           // Increment the actual configured devices, store the state and
           // HW_ID as an numerical value (UINT)
           #statActualConfiguredDevices := #statActualConfiguredDevices + 1;
         ELSE
           ;
         END_IF;

       ELSE
         ; // Device not configured
       END_IF;
     END_FOR;

     #ioSystemData.actualConfiguredDevices := #statActualConfiguredDevices;

     // Mark parameter "Next Device" of the last device in the list
     // --> "Next Device" = negative --> Last device in the list
     #ioSystemData.devices[#statLastDevice].nextDevice := #LAST_DEVICE;

   END_IF; // New IO System detected at input

   #ioSystemData.error := FALSE; // Reset the IO-System error status


   //=============================================================================
   // START DIAGNOSTICS EVALUATION
   //=============================================================================

   //=============================================================================
   // EXISTING DEVICES
   //=============================================================================
   #tempRetValDeviceStates := DeviceStates(LADDR := #ioSystemHwId,
                                           MODE := #MODE_EXIST,
                                           STATE := #statExistingDevices);

   // Check if the block call was successful
   IF (#tempRetValDeviceStates = 0)
   THEN
     // Call ok 
     ;
   ELSIF ((#tempRetValDeviceStates = #ERR_HWID_NOT_EXISTENT)
     OR (#tempRetValDeviceStates = #ERR_LADDR_ADDRESS))
   THEN
     #ioSystemData.error := TRUE;
     #statStatus := INT_TO_WORD(#tempRetValDeviceStates);
     #statStatusID := #ID_DEVICE_STATES_EXISTING;
     #statError := TRUE;
   ELSE
     // Error handling
     #statStatus := INT_TO_WORD(#tempRetValDeviceStates);
     #statStatusID := #ID_DEVICE_STATES_EXISTING;
     #statError := TRUE;
   END_IF;

   //=============================================================================
   // FAULTY DEVICES
   //=============================================================================
   #tempRetValDeviceStates := DeviceStates(LADDR := #ioSystemHwId,
                                           MODE := #MODE_FAULTY,
                                           STATE := #statFaultyDevices);

   // Check if the block call was successful
   IF (#tempRetValDeviceStates = 0)
   THEN
     // Call ok
     ;
   ELSIF ((#tempRetValDeviceStates = #ERR_HWID_NOT_EXISTENT)
     OR (#tempRetValDeviceStates = #ERR_LADDR_ADDRESS))
   THEN
     #ioSystemData.error := TRUE;
     #statStatus := INT_TO_WORD(#tempRetValDeviceStates);
     #statStatusID := #ID_DEVICE_STATES_FAULTY;
     #statError := TRUE;
   ELSE
     // Error handling
     #statStatus := INT_TO_WORD(#tempRetValDeviceStates);
     #statStatusID := #ID_DEVICE_STATES_FAULTY;
     #statError := TRUE;
   END_IF;

   //=============================================================================
   // DISABLED DEVICES
   //=============================================================================
   #tempRetValDeviceStates := DeviceStates(LADDR := #ioSystemHwId,
                                           MODE := #MODE_DISABLED,
                                           STATE := #statDisabledDevices);

   // Check if the block call was successful
   IF (#tempRetValDeviceStates = 0)
   THEN
     // Call ok
     ;
   ELSIF ((#tempRetValDeviceStates = #ERR_HWID_NOT_EXISTENT)
     OR (#tempRetValDeviceStates = #ERR_LADDR_ADDRESS))
   THEN
     #ioSystemData.error := TRUE;
     #statStatus := INT_TO_WORD(#tempRetValDeviceStates);
     #statStatusID := #ID_DEVICE_STATES_DISABLED;
     #statError := TRUE;
   ELSE
     // Error handling
     #statStatus := INT_TO_WORD(#tempRetValDeviceStates);
     #statStatusID := #ID_DEVICE_STATES_DISABLED;
     #statError := TRUE;
   END_IF;

   //=============================================================================
   // PROBLEM DEVICES
   //=============================================================================
   #tempRetValDeviceStates := DeviceStates(LADDR := #ioSystemHwId,
                                           MODE := #MODE_PROBLEM,
                                           STATE := #statProblemDevices);

   // Check if the block call was successful
   IF (#tempRetValDeviceStates = 0)
   THEN
     // Call ok
     ;
   ELSIF ((#tempRetValDeviceStates = #ERR_HWID_NOT_EXISTENT)
     OR (#tempRetValDeviceStates = #ERR_LADDR_ADDRESS))
   THEN
     #ioSystemData.error := TRUE;
     #statStatus := INT_TO_WORD(#tempRetValDeviceStates);
     #statStatusID := #ID_DEVICE_STATES_PROBLEM;
     #statError := TRUE;
   ELSE
     // Error handling
     #statStatus := INT_TO_WORD(#tempRetValDeviceStates);
     #statStatusID := #ID_DEVICE_STATES_PROBLEM;
     #statError := TRUE;
   END_IF;

   //=============================================================================
   // Go through configured devices and check for error
   //=============================================================================
   // Initialize the pointer for the first run 
   #tempDeviceIndex := #ioSystemData.firstDevice;

   WHILE ((#tempDeviceIndex <= "USERDIAG_DEVICES_PER_IO_SYSTEM_UPPER_LIM")
     AND (#tempDeviceIndex > 0))
   DO

     IF (#ioSystemData.devices[#tempDeviceIndex].configured = TRUE)
     THEN

       IF (#statDisabledDevices[#tempDeviceIndex] = TRUE)
       THEN
         //===================
         // Device is disabled
         //===================
         #ioSystemData.devices[#tempDeviceIndex].disabled := TRUE;
         #ioSystemData.devices[#tempDeviceIndex].error := FALSE;
         #ioSystemData.devices[#tempDeviceIndex].faulty := FALSE;
         #ioSystemData.devices[#tempDeviceIndex].problem := FALSE;
         #ioSystemData.devices[#tempDeviceIndex].state := #STATE_DISABLED;

       ELSE
         #ioSystemData.devices[#tempDeviceIndex].disabled := FALSE;

         IF (#statExistingDevices[#tempDeviceIndex] = TRUE)
         THEN
           #ioSystemData.devices[#tempDeviceIndex].exists := TRUE;

           CASE #ioSystemData.devices[#tempDeviceIndex].state OF
             #STATE_WAS_FAULT,
             #STATE_WAS_LOST,
             #STATE_WAS_DISABLED,
             #STATE_PROBLEM_GONE:
               ;
             #STATE_FAULT:
               #ioSystemData.devices[#tempDeviceIndex].state := #STATE_WAS_FAULT;
             #STATE_LOST_CON:
               #ioSystemData.devices[#tempDeviceIndex].state := #STATE_WAS_LOST;
             #STATE_DISABLED:
               #ioSystemData.devices[#tempDeviceIndex].state := #STATE_WAS_DISABLED;
             #STATE_PROBLEM:
               #ioSystemData.devices[#tempDeviceIndex].state := #STATE_PROBLEM_GONE;
             ELSE
               #ioSystemData.devices[#tempDeviceIndex].state := #STATE_OK;
           END_CASE;

         ELSE
           // Device not existent
           #ioSystemData.devices[#tempDeviceIndex].error := TRUE;
           #ioSystemData.error := TRUE; 
           #ioSystemData.devices[#tempDeviceIndex].exists := FALSE;
         END_IF; // End: Device exists


         IF (#statFaultyDevices[#tempDeviceIndex] = FALSE)
         THEN
           // Device is not faulty
           #ioSystemData.devices[#tempDeviceIndex].error := FALSE;
           #ioSystemData.devices[#tempDeviceIndex].faulty := FALSE;

           IF (#statProblemDevices[#tempDeviceIndex] = FALSE)
           THEN
             //============================
             // Device has no problem
             //============================
             #ioSystemData.devices[#tempDeviceIndex].error := FALSE;
             #ioSystemData.devices[#tempDeviceIndex].problem := FALSE;
           ELSE
             //============================
             // Device has a problem
             //============================
             #ioSystemData.devices[#tempDeviceIndex].error := TRUE;
             #ioSystemData.error := TRUE;
             #ioSystemData.devices[#tempDeviceIndex].problem := TRUE;
             #ioSystemData.devices[#tempDeviceIndex].state := #STATE_PROBLEM;
           END_IF;

         ELSE
           // Device is faulty, don't matter what happened
           #ioSystemData.devices[#tempDeviceIndex].error := TRUE;
           #ioSystemData.error := TRUE;
           #ioSystemData.devices[#tempDeviceIndex].faulty := TRUE;

           IF (#statProblemDevices[#tempDeviceIndex] = FALSE)
           THEN
             //============================
             // Device has no problem
             //============================
             #ioSystemData.devices[#tempDeviceIndex].problem := FALSE;
           ELSE
             //============================
             // Device has a problem
             //============================
             #ioSystemData.devices[#tempDeviceIndex].problem := TRUE;
           END_IF;

           IF (#statExistingDevices[#tempDeviceIndex] = FALSE)
           THEN
             //==========================
             // Device is lost
             //==========================
             #ioSystemData.devices[#tempDeviceIndex].state := #STATE_LOST_CON;
             #ioSystemData.devices[#tempDeviceIndex].exists := FALSE;
           ELSE
             //==========================
             // Device is faulty
             //==========================
             #ioSystemData.devices[#tempDeviceIndex].state := #STATE_FAULT;
             #ioSystemData.devices[#tempDeviceIndex].exists := TRUE;
           END_IF;
         END_IF; // End: // Device is not faulty

       END_IF;

       //=============================================================================
       // Set module states
       //=============================================================================
       // Check ModuleStates if device has a problem or is faulty
       IF ((#ioSystemData.devices[#tempDeviceIndex].problem = TRUE)
         OR (#ioSystemData.devices[#tempDeviceIndex].faulty = TRUE))
       THEN

         // PROBLEM MODULE
         #tempRetValModuleStates := ModuleStates(LADDR := #ioSystemData.devices[#tempDeviceIndex].hardwareId,
                                                 MODE := #MODE_PROBLEM,
                                                 STATE := #statDeviceProblemModules);

         // Check if the block call was successful
         IF (#tempRetValModuleStates = 0)
         THEN
           // Call ok 
           ;
         ELSIF ((#tempRetValModuleStates = #ERR_HWID_NOT_EXISTENT)
           OR (#tempRetValModuleStates = #ERR_LADDR_ADDRESS))
         THEN
           #ioSystemData.error := TRUE;
           #statStatus := INT_TO_WORD(#tempRetValModuleStates);
           #statStatusID := #ID_MODULE_STATES_PROBLEM;
           #statError := TRUE;
         ELSE
           // Error handling
           #statStatus := INT_TO_WORD(#tempRetValModuleStates);
           #statStatusID := #ID_MODULE_STATES_PROBLEM;
           #statError := TRUE;
         END_IF;

         // FAULTY MODULE
         #tempRetValModuleStates := ModuleStates(LADDR := #ioSystemData.devices[#tempDeviceIndex].hardwareId,
                                                 MODE := #MODE_FAULTY,
                                                 STATE := #statDeviceFaultyModules);

         // Check if the block call was successful
         IF (#tempRetValModuleStates = 0)
         THEN
           // Call ok 
           ;
         ELSIF ((#tempRetValModuleStates = #ERR_HWID_NOT_EXISTENT)
           OR (#tempRetValModuleStates = #ERR_LADDR_ADDRESS))
         THEN
           #ioSystemData.error := TRUE;
           #statStatus := INT_TO_WORD(#tempRetValModuleStates);
           #statStatusID := #ID_MODULE_STATES_FAULTY;
           #statError := TRUE;
         ELSE
           // Error handling
           #statStatus := INT_TO_WORD(#tempRetValModuleStates);
           #statStatusID := #ID_MODULE_STATES_FAULTY;
           #statError := TRUE;
         END_IF;

         // EXISTING MODULE
         #tempRetValModuleStates := ModuleStates(LADDR := #ioSystemData.devices[#tempDeviceIndex].hardwareId,
                                                 MODE := #MODE_EXIST,
                                                 STATE := #statDeviceExistingModules);

         // Check if the block call was successful
         IF (#tempRetValModuleStates = 0)
         THEN
           // Call ok 
           ;
         ELSIF ((#tempRetValModuleStates = #ERR_HWID_NOT_EXISTENT)
           OR (#tempRetValModuleStates = #ERR_LADDR_ADDRESS))
         THEN
           #ioSystemData.error := TRUE;
           #statStatus := INT_TO_WORD(#tempRetValModuleStates);
           #statStatusID := #ID_MODULE_STATES_EXISTING;
           #statError := TRUE;
         ELSE
           // Error handling
           #statStatus := INT_TO_WORD(#tempRetValModuleStates);
           #statStatusID := #ID_MODULE_STATES_EXISTING;
           #statError := TRUE;
         END_IF;
       END_IF;


       FOR #tempSlotIndex := 0 TO "USERDIAG_SLOTS_PER_DEVICE_UPPER_LIM" DO
         IF (#ioSystemData.devices[#tempDeviceIndex].slots[#tempSlotIndex].configured = TRUE)
         THEN
           CASE #ioSystemData.devices[#tempDeviceIndex].slots[#tempSlotIndex].state OF
             #STATE_WAS_FAULT,
             #STATE_WAS_LOST,
             #STATE_WAS_DISABLED,
             #STATE_PROBLEM_GONE:
               ;
             #STATE_FAULT:
               #ioSystemData.devices[#tempDeviceIndex].slots[#tempSlotIndex].state := #STATE_WAS_FAULT;
             #STATE_LOST_CON:
               #ioSystemData.devices[#tempDeviceIndex].slots[#tempSlotIndex].state := #STATE_WAS_LOST;
             #STATE_DISABLED:
               #ioSystemData.devices[#tempDeviceIndex].slots[#tempSlotIndex].state := #STATE_WAS_DISABLED;
             #STATE_PROBLEM:
               #ioSystemData.devices[#tempDeviceIndex].slots[#tempSlotIndex].state := #STATE_PROBLEM_GONE;
             ELSE
               #ioSystemData.devices[#tempDeviceIndex].slots[#tempSlotIndex].state := #STATE_OK;
           END_CASE;
         END_IF;
       END_FOR;

       CASE #ioSystemData.devices[#tempDeviceIndex].state OF

         #STATE_DISABLED:
           FOR #tempSlotIndex := 0 TO "USERDIAG_SLOTS_PER_DEVICE_UPPER_LIM" DO
             IF (#ioSystemData.devices[#tempDeviceIndex].slots[#tempSlotIndex].configured = TRUE)
             THEN
               //NEW: Set all configured modules of device to disabled
               #ioSystemData.devices[#tempDeviceIndex].slots[#tempSlotIndex].disabled := TRUE;
               #ioSystemData.devices[#tempDeviceIndex].slots[#tempSlotIndex].error := FALSE;
               #ioSystemData.devices[#tempDeviceIndex].slots[#tempSlotIndex].faulty := FALSE;
               #ioSystemData.devices[#tempDeviceIndex].slots[#tempSlotIndex].problem := FALSE;
               #ioSystemData.devices[#tempDeviceIndex].slots[#tempSlotIndex].state := #STATE_DISABLED;
             END_IF;
           END_FOR;

         #STATE_LOST_CON:
           // All modules are faulty when connection is lost
           FOR #tempSlotIndex := 0 TO "USERDIAG_SLOTS_PER_DEVICE_UPPER_LIM" DO
             IF (#ioSystemData.devices[#tempDeviceIndex].slots[#tempSlotIndex].configured = TRUE)
             THEN
               #ioSystemData.devices[#tempDeviceIndex].slots[#tempSlotIndex].error := TRUE;
               #ioSystemData.devices[#tempDeviceIndex].slots[#tempSlotIndex].faulty := TRUE;
               #ioSystemData.devices[#tempDeviceIndex].slots[#tempSlotIndex].problem := TRUE;
               #ioSystemData.devices[#tempDeviceIndex].slots[#tempSlotIndex].exists := FALSE;
               #ioSystemData.devices[#tempDeviceIndex].slots[#tempSlotIndex].state := #STATE_LOST_CON;
             END_IF;
           END_FOR;

         #STATE_FAULT,
         #STATE_PROBLEM:
           // The device is reachable, but faulty because of an error in a
           // subordinated system --> check the modules
           // Store the state of the different module in the diag DB
           FOR #tempSlotIndex := 0 TO "USERDIAG_SLOTS_PER_DEVICE_UPPER_LIM" DO
             IF (#ioSystemData.devices[#tempDeviceIndex].slots[#tempSlotIndex].configured = TRUE)
             THEN
               IF (#statDeviceProblemModules[#tempSlotIndex + 1] = TRUE)
               THEN
                 // Problem in module
                 #ioSystemData.devices[#tempDeviceIndex].slots[#tempSlotIndex].faulty := FALSE;
                 #ioSystemData.devices[#tempDeviceIndex].slots[#tempSlotIndex].error := TRUE;
                 #ioSystemData.devices[#tempDeviceIndex].slots[#tempSlotIndex].problem := TRUE;
                 #ioSystemData.devices[#tempDeviceIndex].slots[#tempSlotIndex].state := #STATE_PROBLEM;

                 IF (#statDeviceFaultyModules[#tempSlotIndex + 1] = TRUE)
                 THEN
                   // Fault in module
                   #ioSystemData.devices[#tempDeviceIndex].slots[#tempSlotIndex].faulty := TRUE;
                   #ioSystemData.devices[#tempDeviceIndex].slots[#tempSlotIndex].state := #STATE_FAULT;
                 END_IF;
               ELSE
                 #ioSystemData.devices[#tempDeviceIndex].slots[#tempSlotIndex].error := FALSE;
                 #ioSystemData.devices[#tempDeviceIndex].slots[#tempSlotIndex].problem := FALSE;
                 #ioSystemData.devices[#tempDeviceIndex].slots[#tempSlotIndex].faulty := FALSE;
               END_IF;

               IF (#statDeviceExistingModules[#tempSlotIndex + 1] = TRUE)
               THEN
                 // Module exists
                 #ioSystemData.devices[#tempDeviceIndex].slots[#tempSlotIndex].exists := TRUE;
               ELSE
                 // Module does not exist
                 #ioSystemData.devices[#tempDeviceIndex].slots[#tempSlotIndex].exists := FALSE;
               END_IF;
             END_IF;
           END_FOR;
         ELSE
           // All modules are okay
           FOR #tempSlotIndex := 0 TO "USERDIAG_SLOTS_PER_DEVICE_UPPER_LIM" DO
             IF (#ioSystemData.devices[#tempDeviceIndex].slots[#tempSlotIndex].configured = TRUE)
             THEN
               #ioSystemData.devices[#tempDeviceIndex].slots[#tempSlotIndex].error := FALSE;
               #ioSystemData.devices[#tempDeviceIndex].slots[#tempSlotIndex].problem := FALSE;
               #ioSystemData.devices[#tempDeviceIndex].slots[#tempSlotIndex].faulty := FALSE;
               #ioSystemData.devices[#tempDeviceIndex].slots[#tempSlotIndex].exists := TRUE;
             END_IF;
           END_FOR;
       END_CASE;
     END_IF;

     // Initialize the pointer for the next run
     #tempDeviceIndex := #ioSystemData.devices[#tempDeviceIndex].nextDevice;
   END_WHILE;


   // Write static values to outputs
   #error := #statError;
   #status := #statStatus;
   #statusID := #statStatusID;
END_FUNCTION_BLOCK

FUNCTION_BLOCK "UserDiag_PLCCheck"   // FB2002, SCL
{ S7_Optimized_Access := 'TRUE' }
VERSION : 0.1
   VAR_INPUT
      plcHwId : Hw_Device;   // Hardware ID
   END_VAR
   VAR_OUTPUT
      error : Bool := FALSE;   // Rising edge informs that an error occurred during the execution of the FB
      status : Word := 16#0000;   // Current status of FB
      statusID : Word;   // Current status ID of calling instruction
   END_VAR
   VAR_IN_OUT
      plcData : "UserDiag_typePLC";   // PLC diagnostics data
   END_VAR
   VAR
      statError : Bool := FALSE;   // Static value for output error
      statStatus : Word := 16#0000;   // Static value for output status
      statStatusID : Word;   // Static value for output statusID
      statGeoAddr : GEOADDR;   // Slot information
      statGeoLaddr : Hw_Any := 16#0000;   // GEO2LOG hardware identifier
      statProblemPlcModulStates : Array[0..#MODULES_STATES_UPPER_LIM] of Bool;   // Storage of the status of all modules in the PLC central station --> State: Problem
      statFaultyPlcModulStates : Array[0..#MODULES_STATES_UPPER_LIM] of Bool;   // Storage of the status of all modules in the PLC central station --> State: Faulty
      statExistingPlcModulStates : Array[0..#MODULES_STATES_UPPER_LIM] of Bool;   // Storage of the status of all modules in the PLC central station --> State: Exists
      statActualCentralModules : USInt := 0;   // Actual number of modules in the central station (PLC)
   END_VAR
   VAR_TEMP
      tempSlotNum : Int;   // Index slot number
      tempRetValGeo : Int;   // GEO2LOG error information
      tempRetValModuleStates : Int;   // Return value system function ModuleStates
   END_VAR
   VAR CONSTANT
      STATUS_EXECUTION_FINISHED : Word := 16#0000;   // Execution finished without errors
      ERR_MAX_SLOTS_PER_PLC : Word := 16#8400;   // There are more modules configured as defined with the user constant: USERDIAG_SLOTS_PER_PLC_UPPER_LIM
      ID_LOCAL : Word := 1;   // StatusID local
      ID_MODULE_STATES_CONFIGURED : Word := 2;   // StatusID during ModuleStates command (configured mode)
      ID_MODULE_STATES_FAULTY : Word := 3;   // StatusID during ModuleStates command (faulty mode)
      ID_MODULE_STATES_PROBLEM : Word := 4;   // StatusID during ModuleStates command (problem mode)
      ID_MODULE_STATES_EXISTING : Word := 5;   // StatusID during ModuleStates command (existing mode)
      ID_LED : Word := 12;   // StatusID occurred during LED command
      MODE_FAULTY : USInt := 2;   // Used for instruction DeviceStates, read out all faulty devices
      MODE_EXIST : USInt := 4;   // Used for instruction DeviceStates, read out all devices not reachable
      MODE_PROBLEM : USInt := 5;   // Used for instruction DeviceStates, read out all devices with several problems
      STATE_OK : USInt := 1;   // Module state: ok
      STATE_FAULT : USInt := 2;   // Modulestate: fault
      STATE_PROBLEM : USInt := 5;   // Module state: problem
      STATE_WAS_FAULT : USInt := 12;   // Module state: was fault
      STATE_PROBLEM_GONE : USInt := 15;   // Module state: had a problem
      MODULE_OF_PLC : USInt := 4;   // GEO2LOG structure: HW type = 4
      CPU : USInt := 0;   // GEO2LOG structure: Area = 0
      CENTRAL_SYSTEM : USInt := 0;   // GEO2LOG structure: IO System = 0
      CENTRAL_STATION : USInt := 0;   // GEO2LOG structure: Station = 0
      NO_LED : Int := 0;   // LED does not exist
      LED_OFF : Int := 1;   // LED is permanently switched off
      LED_NO_INFO : Int := 9;   // LED exists, but status information not available
      MODULES_STATES_UPPER_LIM : Int := 127;   // Upper array limit for output tag of instruction ModuleStates
      ERROR_LED : UInt := 2;   // Identification number of the LED
   END_VAR
BEGIN
   //=============================================================================
   //SIEMENS AG
   //(c)Copyright 2017 All Rights Reserved
   //-----------------------------------------------------------------------------
   //Library: 
   //Tested with: S7-1516-3 PN/DP FW 2.5
   //Engineering: TIA Portal V14 Update1
   //Restrictions: Call in cyclic OB
   //Requirements: -
   //Functionality: Determine plc state and local module states
   //-----------------------------------------------------------------------------
   //Change log table:
   //Version  Date       Expert in charge                Changes applied
   //01.00.00 27.01.2017 Siemens Industry Online Support First released version
   //01.00.01 20.12.2017 Siemens Industry Online Support actualConfiguredSlots >= 1
   //01.00.02 27.02.2018 Siemens Industry Online Support Minor corrections
   //=============================================================================

   IF (#plcData.hardwareId = 0)
   THEN
     #statGeoAddr.HWTYPE := #MODULE_OF_PLC;      // Hardware type 4: module
     #statGeoAddr.AREA := #CPU;                  // Area ID 0: CPU
     #statGeoAddr.IOSYSTEM := #CENTRAL_SYSTEM;   // PROFINET IO system (0 = central unit in the rack)
     #statGeoAddr.STATION := #CENTRAL_STATION;   // Number of the rack if area identifier AREA = 0 (central module)

     #statStatus := #STATUS_EXECUTION_FINISHED;
     #statStatusID := 0;
     #statError := FALSE;
     #statActualCentralModules := 0;

     FOR #tempSlotNum := 0 TO "USERDIAG_SLOTS_PER_PLC_UPPER_LIM" DO
       // Slot number
       #statGeoAddr.SLOT := INT_TO_UINT(#tempSlotNum);
       // read LADDR from local modules
       #tempRetValGeo := GEO2LOG(GEOADDR := #statGeoAddr,
                                 LADDR => #statGeoLaddr);
       // Check Retval
       IF ((#tempRetValGeo = 0)
         AND (#statGeoLaddr <> 16#0))
       THEN
         // Store LADDR from local modules in diagnostic data block
         IF (#tempSlotNum = 1)
         THEN
           #plcData.hardwareId := #statGeoLaddr;
         END_IF;
         #plcData.slots[#tempSlotNum].hardwareId := #statGeoLaddr;
         #statActualCentralModules := #statActualCentralModules + 1;
         #plcData.slots[#tempSlotNum].configured := TRUE;
       ELSE
         // If the return value ist not = 0 --> the device/system/module is not
         // configured --> No error handling
         // set LADDR from local modules to 0 in diagnostic data block
         #plcData.slots[#tempSlotNum].hardwareId := 0;
         #plcData.slots[#tempSlotNum].configured := FALSE;
       END_IF;
       // Store the actual configured devices in the diagnostics DB
       #plcData.actualConfiguredSlots := #statActualCentralModules;
     END_FOR;

     // Check if further slots are configured
     #statGeoAddr.SLOT := INT_TO_UINT(#tempSlotNum);

     #tempRetValGeo := GEO2LOG(GEOADDR := #statGeoAddr,
                               LADDR => #statGeoLaddr);

     IF ((#tempRetValGeo = 0)
       AND (#statGeoLaddr <> 16#0))
     THEN
       // In the PLC are more slots configured as defined with the user constant
       #statStatus := #ERR_MAX_SLOTS_PER_PLC;
       #statStatusID := #ID_LOCAL;
       #statError := TRUE;
     END_IF;

   END_IF;

   // Reset PLC error state
   #plcData.error := FALSE;

   //=============================================================================
   // Check modul states from LOCAL MODULES
   //=============================================================================
   // Check if central module are available - at least one module is always
   // configured, the PLC itself
   IF (#plcData.actualConfiguredSlots >= 1)
   THEN

     // Check the status of the local modules
     #tempRetValModuleStates := ModuleStates(LADDR := #plcHwId,
                                             MODE := #MODE_PROBLEM,
                                             STATE := #statProblemPlcModulStates);

     // Check if the block call was successful
     IF (#tempRetValModuleStates <> 0)
     THEN
       // Error handling
       #statStatus := INT_TO_WORD(#tempRetValModuleStates);
       #statStatusID := #ID_MODULE_STATES_PROBLEM;
       #statError := TRUE;
     ELSE
       ; // Everything is ok!
     END_IF;

     #tempRetValModuleStates := ModuleStates(LADDR := #plcHwId,
                                             MODE := #MODE_FAULTY,
                                             STATE := #statFaultyPlcModulStates);

     // Check if the block call was successful
     IF (#tempRetValModuleStates <> 0)
     THEN
       // Error handling
       #statStatus := INT_TO_WORD(#tempRetValModuleStates);
       #statStatusID := #ID_MODULE_STATES_FAULTY;
       #statError := TRUE;
     ELSE
       ; // Everything is ok!
     END_IF;

     #tempRetValModuleStates := ModuleStates(LADDR := #plcHwId,
                                             MODE := #MODE_EXIST,
                                             STATE := #statExistingPlcModulStates);

     // Check if the block call was successful
     IF (#tempRetValModuleStates <> 0)
     THEN
       // Error handling
       #statStatus := INT_TO_WORD(#tempRetValModuleStates);
       #statStatusID := #ID_MODULE_STATES_EXISTING;
       #statError := TRUE;
     ELSE
       ; // Everything is ok!
     END_IF;

   ELSE
     ; // There are no central moduls configured
   END_IF;

   //=============================================================================
   // Set module states of LOCAL MODULES
   //=============================================================================
   #tempSlotNum := 0;
   WHILE (#tempSlotNum <= #plcData.actualConfiguredSlots)
   DO
     IF (#plcData.slots[#tempSlotNum].configured)
     THEN
       IF (#statExistingPlcModulStates[#tempSlotNum + 1] = TRUE)
       THEN
         #plcData.slots[#tempSlotNum].exists := TRUE;
         CASE #plcData.slots[#tempSlotNum].state OF
           #STATE_WAS_FAULT,
           #STATE_PROBLEM_GONE:
             ;
           #STATE_FAULT:
             #plcData.slots[#tempSlotNum].state := #STATE_WAS_FAULT;
           #STATE_PROBLEM:
             #plcData.slots[#tempSlotNum].state := #STATE_PROBLEM_GONE;
           ELSE
             #plcData.slots[#tempSlotNum].state := #STATE_OK;
         END_CASE;
       ELSE
         #plcData.slots[#tempSlotNum].error := TRUE;
         #plcData.error := TRUE;
         #plcData.slots[#tempSlotNum].exists := FALSE;
       END_IF;

       IF (#statFaultyPlcModulStates[#tempSlotNum + 1] = TRUE)
       THEN
         // Modul is faulty
         #plcData.slots[#tempSlotNum].faulty := TRUE;
         #plcData.slots[#tempSlotNum].problem := TRUE;
         #plcData.slots[#tempSlotNum].error := TRUE;
         #plcData.slots[#tempSlotNum].state := #STATE_FAULT;
       ELSIF (#statProblemPlcModulStates[#tempSlotNum + 1] = TRUE)
       THEN
         // Modul has a problem
         #plcData.slots[#tempSlotNum].faulty := FALSE;
         #plcData.slots[#tempSlotNum].problem := TRUE;
         #plcData.slots[#tempSlotNum].error := TRUE;
         #plcData.slots[#tempSlotNum].state := #STATE_PROBLEM;
       ELSE
         // Modul is OK
         #plcData.slots[#tempSlotNum].error := FALSE;
         #plcData.slots[#tempSlotNum].problem := FALSE;
         #plcData.slots[#tempSlotNum].faulty := FALSE;
       END_IF;

       // Error in PLC - Slot = 1, but index must be increased by 1, because of bit 0 = group display
       // --> used index = 2
       IF (#statProblemPlcModulStates[2] = TRUE)
         OR (#statFaultyPlcModulStates[2] = TRUE)
       THEN
         #plcData.error := TRUE;
       END_IF;
     END_IF;

     #tempSlotNum := #tempSlotNum + 1;
   END_WHILE;

   // Write static values to outputs
   #error := #statError;
   #status := #statStatus;
   #statusID := #statStatusID;

   //----------------------------------------------------------------------------------------------
END_FUNCTION_BLOCK

FUNCTION_BLOCK "UserDiag_Diagnostics"   // FB2003, LAD
{ S7_Optimized_Access := 'TRUE' }
VERSION : 0.1
// //============================================================================
// //SIEMENS AG
// //(c)Copyright 2017 All Rights Reserved
// //-----------------------------------------------------------------------------
// //Library: -
// //Tested with: S7-1516-3 PN/DP FW 2.5
// //Engineering: TIA Portal V14 Update1
// //Restrictions: -
// //Requirements: -
// //Functionality: Main FB for diagnostics
// //-----------------------------------------------------------------------------
// //Change log table:
// //Version  Date              Expert in charge                               Changes applied
// //01.00.00 25.04.2017 Siemens Industry Online Support First released version
// //01.01.00 01.12.2017 Siemens Industry Online Support Renamed in "UserDiag_Diagnostics"
// //                                                                                                    Check Flag "startDiag"
// //============================================================================
   VAR_IN_OUT
      startDiag : Bool;   // Startflag for diagnostic
      plcData : "UserDiag_typePLC";   // PLC diagnostics data
      ioSystemData : Array[1.."USERDIAG_IO_SYSTEMS_UPPER_LIM"] of "UserDiag_typeIOSystem";   // IO-System diagnostics data
   END_VAR
   VAR
      instPLCCheck : "UserDiag_PLCCheck";   // Instance of "UserDiag_PLCCheck"
      instIOSystemCheck1 : "UserDiag_IOSystemCheck";   // Instance of "UserDiag_IOSystemCheck"
      instIOSystemCheck2 : "UserDiag_IOSystemCheck";   // Instance of "UserDiag_IOSystemCheck"
   END_VAR
BEGIN

REGION Network 1: Check Startflag for diagnostic
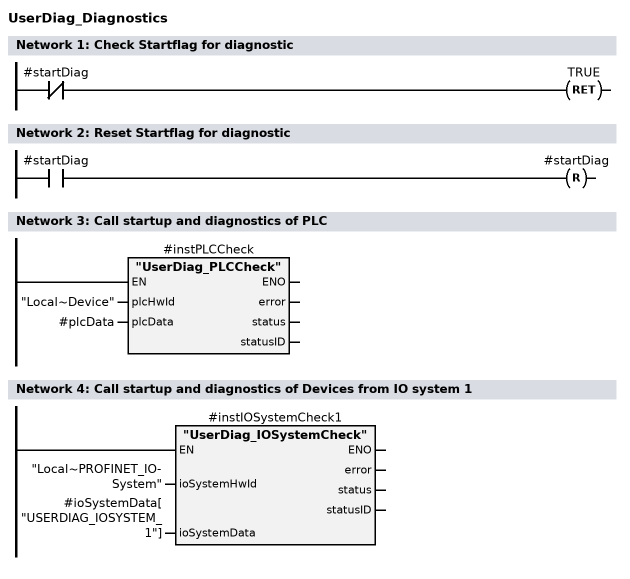
   IF NOT #startDiag THEN
       ENO := TRUE;
       RETURN;
   END_IF;
END_REGION

REGION Network 2: Reset Startflag for diagnostic
   RUNG wire#powerrail
      Contact( #startDiag )
      R_Coil( #startDiag )
   END_RUNG
   // the same network as SCL:
   IF #startDiag THEN #startDiag := FALSE; END_IF;
END_REGION

REGION Network 3: Call startup and diagnostics of PLC
   RUNG wire#powerrail
      #instPLCCheck(plcHwId := "Local~Device", plcData := #plcData, error =>, status =>, statusID =>)
   END_RUNG
   // the same network as SCL:
   #instPLCCheck(plcHwId := "Local~Device", plcData := #plcData);   // "UserDiag_PLCCheck"
END_REGION

REGION Network 4: Call startup and diagnostics of Devices from IO system 1
   RUNG wire#powerrail
      #instIOSystemCheck1(ioSystemHwId := "Local~PROFINET_IO-System", ioSystemData := #ioSystemData["USERDIAG_IOSYSTEM_1"], error =>, status =>, statusID =>)
   END_RUNG
   // the same network as SCL:
   #instIOSystemCheck1(ioSystemHwId := "Local~PROFINET_IO-System",   // "UserDiag_IOSystemCheck"
                       ioSystemData := #ioSystemData["USERDIAG_IOSYSTEM_1"]);
END_REGION
END_FUNCTION_BLOCK

FUNCTION_BLOCK "UserDiag_GetIPAddress"   // FB2005, SCL
{ S7_Optimized_Access := 'TRUE' }
VERSION : 0.1
   VAR_OUTPUT
      error : Bool := FALSE;   // Rising edge informs that an error occurred during the execution of the FB
      status : Word := 16#0000;   // Current status of FB
      statusID : Word;   // Current status ID of calling instruction
   END_VAR
   VAR_IN_OUT
      ioSystemData : "UserDiag_typeIOSystem";   // IO-System diagnostics data
   END_VAR
   VAR
      statError : Bool := FALSE;   // Static value for output error
      statStatus : Word := 16#0000;   // Static value for output status
      statStatusID : Word;   // Static value for output statusID
      instGetStationInfo : GetStationInfo;   // Instance of GetStationInfo
      statFirstDeviceFlag : Bool := TRUE;   // Help tag for the first device in the linked list
      statDeviceIndex : Int;   // Device/slave index
   END_VAR
   VAR_TEMP
      tempIP : IF_CONF_v4;   // Temporary IP address
   END_VAR
   VAR CONSTANT
      STATUS_EXECUTION_FINISHED : Word := 16#0000;   // Execution finished without errors
      ID_GET_STATION_INFO : Word := 12;   // StatusID during GetStationInfo command
      MODE_IPV4 : UInt := 1;   // Address parameter according to IPv4
      LAST_DEVICE : Int := -1;   // No next device
   END_VAR
BEGIN
   //=============================================================================
   //SIEMENS AG
   //(c)Copyright 2015 All Rights Reserved
   //-----------------------------------------------------------------------------
   //Library: 
   //Tested with: S7-1516-3 PN/DP FW 2.5
   //Engineering: TIA Portal V14 Update1
   //Restrictions: Call in cyclic OB
   //Requirements: -
   //Functionality: Get IP address of IO devices
   //-----------------------------------------------------------------------------
   //Change log table:
   //Version  Date       Expert in charge                Changes applied
   //01.00.00 20.12.2017 Siemens Industry Online Support First released version
   //=============================================================================

   //=============================================================================
   // Go through existing devices and get IP address
   //=============================================================================
   // Initialize the pointer for the first run 
   IF (#statFirstDeviceFlag = TRUE)
   THEN
     #statDeviceIndex := #ioSystemData.firstDevice;
     #statFirstDeviceFlag := FALSE;
   END_IF;

   // Check and store the IP address, if the device is existing
   // GetStationInfo is an acyclic instruction. In the FB, the
   // instruction has to be repeated until it is done or error
   IF ((#ioSystemData.number >= 100)
     AND (#ioSystemData.number <= 115)
     AND (#ioSystemData.devices[#statDeviceIndex].exists = TRUE)
     AND (#ioSystemData.devices[#statDeviceIndex].ipAddress.ADDR[1] = 0))
   THEN
     // Get IP address of each decive in PN System
     #instGetStationInfo(REQ := TRUE,
                         LADDR := #ioSystemData.devices[#statDeviceIndex].hardwareId,
                         MODE := #MODE_IPV4,
                         DATA := #tempIP);

     IF (#instGetStationInfo.ERROR = TRUE)
     THEN
       // Error handling
       #statStatus := #instGetStationInfo.STATUS;
       #statStatusID := #ID_GET_STATION_INFO;
       #statError := TRUE;

       // Everything is ok --> Copy IP address    
     ELSIF (#instGetStationInfo.DONE = TRUE)
     THEN
       #ioSystemData.devices[#statDeviceIndex].ipAddress := #tempIP.InterfaceAddress;

       // Initialize the pointer for the next run
       #statDeviceIndex := #ioSystemData.devices[#statDeviceIndex].nextDevice;
     ELSE
       ;
     END_IF;
   ELSE
     // Initialize the pointer for the next run
     #statDeviceIndex := #ioSystemData.devices[#statDeviceIndex].nextDevice;
   END_IF;

   // Check last device
   IF (#statDeviceIndex = #LAST_DEVICE)
   THEN
     #statDeviceIndex := #ioSystemData.firstDevice;
   END_IF;

   // Write static values to outputs
   #error := #statError;
   #status := #statStatus;
   #statusID := #statStatusID;
END_FUNCTION_BLOCK

FUNCTION_BLOCK "UserDiag_DiagnosticsHmi"   // FB2006, SCL
{ S7_Optimized_Access := 'TRUE' }
VERSION : 0.1
   VAR_IN_OUT
      plcData : "UserDiag_typePLC";   // PLC diagnostics data
      ioSystemData : Array[1.."USERDIAG_IO_SYSTEMS_UPPER_LIM"] of "UserDiag_typeIOSystem";   // IO-System diagnostics data
      hmiData : "UserDiag_typeHmiData";   // HMI data
   END_VAR
   VAR
      statFirstRun : Bool := TRUE;   // TRUE after startup
      instAckTON : TON_TIME;   // Instance of TON_TIME for auto acknowledge
      instRisFilterErrorDevices : R_TRIG;   // Instance of R_TRIG for filter error devices
      statActIOSystem : Int;   // Actual IO system
      statActScreenDevices : Int;   // Actual screen devices
      statActDeviceOfScreen : Int;   // Actual device of screen
   END_VAR
   VAR_TEMP
      tempIndex : Int;   // Index of configured devices/slaves
      tempDeviceIndex : Int;   // Device/slave index
      tempDeviceCount : Int;   // Device counter
      tempSlotIndex : Int;   // Slot index
      tempIoIndex : Int;   // IO system index
      tempErrorStateLower : Bool;   // Temp error at lower screen
      tempErrorStateUpper : Bool;   // Temp error at upper screen
   END_VAR
   VAR CONSTANT
      STATE_OK : USInt := 1;   // Device/module state: ok
      STATE_FAULT : USInt := 2;   // Device/modul state: fault
      STATE_LOST_CON : USInt := 3;   // Device/modul state: lost connection
      STATE_DISABLED : USInt := 4;   // Device/modul state: disabled
      STATE_PROBLEM : USInt := 5;   // Device/modul state: problem
      STATE_WAS_FAULT : USInt := 12;   // Device/module state: was fault
      STATE_WAS_LOST : USInt := 13;   // Device/module state: connection was lost
      STATE_WAS_DISABLED : USInt := 14;   // Device/module state: device was disabled
      STATE_PROBLEM_GONE : USInt := 15;   // Device/module state: had a problem
   END_VAR
BEGIN
   //=============================================================================
   //SIEMENS AG
   //(c)Copyright 2017 All Rights Reserved
   //-----------------------------------------------------------------------------
   //Library: 
   //Tested with: S7-1516-3 PN FW 2.5
   //Engineering: TIA Portal V14 Update1
   //Restrictions: Call in cyclic OB
   //Requirements: -
   //Functionality: Copy and control diagnostics information for visualization
   //-----------------------------------------------------------------------------
   //Change log table:
   //Version  Date       Expert in charge                Changes applied
   //01.00.00 27.01.2017 Siemens Industry Online Support First released version
   //01.01.00 17.10.2017 Siemens Industry Online Support Single parameters 
   //                                                    replaced by "hmiData"
   //01.02.00 20.12.2017 Siemens Industry Online Support Static tags for consistence
   //                                                    (Bereichslängenfehler)
   //=============================================================================

   //=============================================================================
   // Auto acknowledge after waiting time
   //=============================================================================
   #instAckTON(IN := #statFirstRun,
               PT := INT_TO_TIME(#hmiData.ackWaitTime * 1000));

   IF (#instAckTON.Q = TRUE)
   THEN
     // Acknowledge IO systems
     FOR #tempIoIndex := 1 TO "USERDIAG_IO_SYSTEMS_UPPER_LIM" DO
       // Initialize the pointer for the first run 
       #tempDeviceIndex := #ioSystemData[#tempIoIndex].firstDevice;

       WHILE ((#tempDeviceIndex <= "USERDIAG_DEVICES_PER_IO_SYSTEM_UPPER_LIM")
         AND (#tempDeviceIndex > 0))
       DO
         IF (#ioSystemData[#tempIoIndex].devices[#tempDeviceIndex].configured = TRUE)
         THEN
           // Acknowledge "was diabled/faulty/prolem/lost state"
           IF ((#ioSystemData[#tempIoIndex].devices[#tempDeviceIndex].state = #STATE_WAS_DISABLED)
             OR (#ioSystemData[#tempIoIndex].devices[#tempDeviceIndex].state = #STATE_WAS_FAULT)
             OR (#ioSystemData[#tempIoIndex].devices[#tempDeviceIndex].state = #STATE_WAS_LOST)
             OR (#ioSystemData[#tempIoIndex].devices[#tempDeviceIndex].state = #STATE_PROBLEM_GONE))
           THEN
             // Device
             #ioSystemData[#tempIoIndex].devices[#tempDeviceIndex].state := #STATE_OK;
             // Modules
             FOR #tempSlotIndex := 0 TO "USERDIAG_SLOTS_PER_DEVICE_UPPER_LIM" DO
               IF (#ioSystemData[#tempIoIndex].devices[#tempDeviceIndex].slots[#tempSlotIndex].configured = TRUE)
               THEN
                 #ioSystemData[#tempIoIndex].devices[#tempDeviceIndex].slots[#tempSlotIndex].state := #STATE_OK;
               END_IF;
             END_FOR;
           END_IF;
         END_IF;
         // Initialize the pointer for the next run
         #tempDeviceIndex := #ioSystemData[#tempIoIndex].devices[#tempDeviceIndex].nextDevice;
       END_WHILE;

       // Acknowledge local modules
       FOR #tempIndex := 0 TO "USERDIAG_SLOTS_PER_PLC_UPPER_LIM" DO
         IF ((#plcData.slots[#tempIndex].state = #STATE_WAS_FAULT)
           OR (#plcData.slots[#tempIndex].state = #STATE_PROBLEM_GONE))
         THEN
           #plcData.slots[#tempIndex].state := #STATE_OK;
         END_IF;
       END_FOR;
     END_FOR;

     #statFirstRun := FALSE;
   END_IF;

   //=============================================================================
   // Check if a IO system is selected
   //=============================================================================
   // Copy to static tags for consistence
   #statActIOSystem := #hmiData.actIOSystem;
   #statActScreenDevices := #hmiData.actScreenDevices;
   #statActDeviceOfScreen := #hmiData.actDeviceOfScreen;

   IF ((#statActIOSystem >= 1)
     AND (#statActIOSystem <= "USERDIAG_IO_SYSTEMS_UPPER_LIM"))
   THEN
     #hmiData.actIOSystemData.actIOSystemNumber := UINT_TO_INT(#ioSystemData[#statActIOSystem].number);

     // Calculate the maximum count of screens to visualize the devices/slaves
     #hmiData.maxScreensDevices := 1;

     IF ((#ioSystemData[#statActIOSystem].actualConfiguredDevices MOD "USERDIAG_DEVICES_PER_SCREEN_UPPER_LIM") = 0)
     THEN
       #hmiData.maxScreensDevices := #ioSystemData[#statActIOSystem].actualConfiguredDevices / "USERDIAG_DEVICES_PER_SCREEN_UPPER_LIM";
     ELSE
       #hmiData.maxScreensDevices := #ioSystemData[#statActIOSystem].actualConfiguredDevices / "USERDIAG_DEVICES_PER_SCREEN_UPPER_LIM" + 1;
     END_IF;

     //=============================================================================
     // Acknowledge
     //=============================================================================
     IF (#hmiData.ackStates = TRUE)
     THEN
       // Initialize the pointer for the first run 
       #tempDeviceIndex := #ioSystemData[#statActIOSystem].firstDevice;

       WHILE ((#tempDeviceIndex <= "USERDIAG_DEVICES_PER_IO_SYSTEM_UPPER_LIM")
         AND (#tempDeviceIndex > 0))
       DO
         IF (#ioSystemData[#statActIOSystem].devices[#tempDeviceIndex].configured = TRUE)
         THEN
           // Acknowledge "was diabled/faulty/prolem/lost state"
           IF ((#ioSystemData[#statActIOSystem].devices[#tempDeviceIndex].state = #STATE_WAS_DISABLED)
             OR (#ioSystemData[#statActIOSystem].devices[#tempDeviceIndex].state = #STATE_WAS_FAULT)
             OR (#ioSystemData[#statActIOSystem].devices[#tempDeviceIndex].state = #STATE_WAS_LOST)
             OR (#ioSystemData[#statActIOSystem].devices[#tempDeviceIndex].state = #STATE_PROBLEM_GONE))
           THEN
             // Device
             #ioSystemData[#statActIOSystem].devices[#tempDeviceIndex].state := #STATE_OK;
             // Modules
             FOR #tempSlotIndex := 0 TO "USERDIAG_SLOTS_PER_DEVICE_UPPER_LIM" DO
               IF (#ioSystemData[#statActIOSystem].devices[#tempDeviceIndex].slots[#tempSlotIndex].configured = TRUE)
               THEN
                 #ioSystemData[#statActIOSystem].devices[#tempDeviceIndex].slots[#tempSlotIndex].state := #STATE_OK;
               END_IF;
             END_FOR;
           END_IF;
         END_IF;
         // Initialize the pointer for the next run
         #tempDeviceIndex := #ioSystemData[#statActIOSystem].devices[#tempDeviceIndex].nextDevice;
       END_WHILE;
     END_IF;

     //=============================================================================
     // Copy number and status to HMI array
     //=============================================================================
     // Initialize the pointer for the first run 
     #tempDeviceIndex := #ioSystemData[#statActIOSystem].firstDevice;
     // Initialize the pointer for devices on screen
     #tempIndex := 1;
     #tempDeviceCount := 0;

     #instRisFilterErrorDevices(CLK := #hmiData.filterErrorDevices);
     IF (#instRisFilterErrorDevices.Q = TRUE)
     THEN
       #statActScreenDevices := 1;
     END_IF;

     WHILE ((#tempDeviceIndex <= "USERDIAG_DEVICES_PER_IO_SYSTEM_UPPER_LIM")
       AND (#tempDeviceIndex > 0)
       AND (#tempIndex <= "USERDIAG_DEVICES_PER_SCREEN_UPPER_LIM"))
     DO
       IF (#hmiData.filterErrorDevices = FALSE)
       THEN
         IF (#ioSystemData[#statActIOSystem].devices[#tempDeviceIndex].configured = TRUE)
         THEN
           #tempDeviceCount := #tempDeviceCount + 1;

           IF ((#tempDeviceCount > ((#statActScreenDevices - 1) * "USERDIAG_DEVICES_PER_SCREEN_UPPER_LIM"))
             AND (#tempDeviceCount <= (#statActScreenDevices * "USERDIAG_DEVICES_PER_SCREEN_UPPER_LIM")))
           THEN
             // Device configured, status can be copied
             #hmiData.actIOSystemData.actIODeviceNumbers[#tempIndex] := #ioSystemData[#statActIOSystem].devices[#tempDeviceIndex].number;
             #hmiData.actIOSystemData.actIODeviceState[#tempIndex] := #ioSystemData[#statActIOSystem].devices[#tempDeviceIndex].state;
             // Increment index of device per screen
             #tempIndex := #tempIndex + 1;

           END_IF;
         END_IF;
         // Initialize the pointer for the next run
         #tempDeviceIndex := #ioSystemData[#statActIOSystem].devices[#tempDeviceIndex].nextDevice;

         //=============================================================================
         // If filter is enabled, copy number and status of faulty devices to HMI array
         //=============================================================================
       ELSIF (#hmiData.filterErrorDevices = TRUE)
       THEN
         IF ((#ioSystemData[#statActIOSystem].devices[#tempDeviceIndex].configured = TRUE)
           AND (#ioSystemData[#statActIOSystem].devices[#tempDeviceIndex].state > 1))
         THEN
           #tempDeviceCount := #tempDeviceCount + 1;

           IF ((#tempDeviceCount > ((#statActScreenDevices - 1) * "USERDIAG_DEVICES_PER_SCREEN_UPPER_LIM"))
             AND (#tempDeviceCount <= (#statActScreenDevices * "USERDIAG_DEVICES_PER_SCREEN_UPPER_LIM")))
           THEN
             // Device configured, status can be copied
             #hmiData.actIOSystemData.actIODeviceNumbers[#tempIndex] := #ioSystemData[#statActIOSystem].devices[#tempDeviceIndex].number;
             #hmiData.actIOSystemData.actIODeviceState[#tempIndex] := #ioSystemData[#statActIOSystem].devices[#tempDeviceIndex].state;
             // Increment index of device per screen
             #tempIndex := #tempIndex + 1;

           END_IF;
         END_IF;
         // Initialize the pointer for the next run
         #tempDeviceIndex := #ioSystemData[#statActIOSystem].devices[#tempDeviceIndex].nextDevice;

       END_IF;
     END_WHILE;

     // clear screen
     FOR #tempIndex := #tempIndex TO "USERDIAG_DEVICES_PER_SCREEN_UPPER_LIM" DO
       // No device configured
       #hmiData.actIOSystemData.actIODeviceNumbers[#tempIndex] := 0;
       #hmiData.actIOSystemData.actIODeviceState[#tempIndex] := 0;
     END_FOR;